// TIA Portal project "TESTV18" (V18) (continued)
REGION Network 8: HMI Command
   RUNG wire#powerrail
      Contact( "DB_AUX".HMI_Bit.HMIb5 )
      Coil( "DB_AUX".AXIS1.PLCToPCON.CTRL2.CTRL2_Sig_SON )
   END_RUNG
   RUNG wire#powerrail
      Contact( "DB_AUX".HMI_Bit.HMIb6 )
      Coil( "DB_AUX".AXIS1.PLCToPCON.CTRL2.CTRL2_Sig_DSTR )
   END_RUNG
   RUNG wire#powerrail
      Contact( "DB_AUX".HMI_Bit.HMIb7 )
      Coil( "DB_AUX".AXIS1.PLCToPCON.CTRL2.CTRL2_Sig_HOME )
   END_RUNG
   RUNG wire#powerrail
      Contact( "DB_AUX".HMI_Bit.HMIb8 )
      Coil( "DB_AUX".AXIS1.PLCToPCON.CTRL2."CTRL2_Sig_JOG+" )
   END_RUNG
   RUNG wire#powerrail
      Contact( "DB_AUX".HMI_Bit.HMIb9 )
      Coil( "DB_AUX".AXIS1.PLCToPCON.CTRL2."CTRL2_Sig_JOG-" )
   END_RUNG
   RUNG wire#powerrail
      Contact( "DB_AUX".HMI_Bit.HMIb10 )
      Coil( "DB_AUX".AXIS1.PLCToPCON.CTRL2.CTRL2_Sig_RES )
   END_RUNG
   // the same network as SCL:
   "DB_AUX".AXIS1.PLCToPCON.CTRL2.CTRL2_Sig_SON := "DB_AUX".HMI_Bit.HMIb5;
   "DB_AUX".AXIS1.PLCToPCON.CTRL2.CTRL2_Sig_DSTR := "DB_AUX".HMI_Bit.HMIb6;
   "DB_AUX".AXIS1.PLCToPCON.CTRL2.CTRL2_Sig_HOME := "DB_AUX".HMI_Bit.HMIb7;
   "DB_AUX".AXIS1.PLCToPCON.CTRL2."CTRL2_Sig_JOG+" := "DB_AUX".HMI_Bit.HMIb8;
   "DB_AUX".AXIS1.PLCToPCON.CTRL2."CTRL2_Sig_JOG-" := "DB_AUX".HMI_Bit.HMIb9;
   "DB_AUX".AXIS1.PLCToPCON.CTRL2.CTRL2_Sig_RES := "DB_AUX".HMI_Bit.HMIb10;
END_REGION
END_ORGANIZATION_BLOCK

// folder: LIBRERIE OPEN/0 Bit logic operations

FUNCTION "LGF_BitToggle" : DWord   // FC10033, SCL
TITLE = LGF_BitToggle
{ S7_Optimized_Access := 'TRUE' }
AUTHOR : Siemens_SIMATIC_Systems_Support
FAMILY : LGF
NAME : LGF_BitToggle
// Dieser Baustein toggelt (von TRUE nach FALSE und umgekehrt) ein Bit an vorgegebener Stelle in einer Variablen vom Datentyp DWORD.    
// Anstelle von DWord kann auch Word und Byte verwendet werden, indem der übergebene Parameter mit z. B. BYTE_TO_DWORD und das Ergebnis mit DWORD_TO_BYTE konvertiert wird.
// This block toggles (from TRUE to FALSE and vice versa) a bit at a predefined position in a variable of the data type DWORD.  
// Alternatively, Word and Byte can be used instead of DWord by converting the passed parameter with, for example, BYTE_TO_DWORD and the result with DWORD_TO_BYTE
   VAR_INPUT
      value : DWord;   // Tag where the bit has to be toggled / Variable, an der das Bit getoggelt wird.
      bitNo : USInt;   // Bit number to be toggled in the “value” parameter. / Bitnummer, die im Parameter "value" getoggelt werden soll.
   END_VAR
   // Ret_Val : Tag with toggled bit / Variable mit getoggeltem Bit.
   VAR CONSTANT
      TRUE_BOOL_BIT : DWord := 16#0001;   // Just one bit which is true, to shift in Dword for masking / Ein einzelnes Bit mit Wert := TRUE zum schieben im Dword und zur Maskierung
      MAX_NO_OF_BITS : USInt := 32;   // Maximum bits in a DWord = 32 / Maximalanzahl an Bits in einem Dword = 32
   END_VAR
BEGIN
   REGION BLOCK INFO HEADER
     //===============================================================================
     // SIEMENS AG / (c)Copyright 2019
     //-------------------------------------------------------------------------------
     // Title:            LGF_BitToggle
     // Comment/Function: Toggle bit in elementary datatype - DWord
     //                   can be used for Word and Byte as well, by convert
     //                   the passed paramter and the result using for e.g. Dword_to_Byte
     // Library/Family:   LGF (Library General Functions)
     // Author:           Siemens Digital Industry
     // Tested with:      CPU1212C DC/DC/DC FW:V4.2
     // Engineering:      TIA Portal V15.1
     // Restrictions:     ENO not in use, set to true, no error handling
     // Requirements:     PLC (S7-1200 / S7-1500)
     //-------------------------------------------------------------------------------
     // Change log table:
     // Version  | Date       | Expert in charge         | Changes applied
     // 01.00.00 | 06.06.2015 | Siemens Industry Support | first release
     // 03.00.00 | 23.04.2020 | Siemens Industry Support | Set version to V3.0.0
     //                         harmonize the version of the whole library
     // 03.00.01 | 19.01.2021 | Simatic Systems Support
     //                         Insert documentation
     //===============================================================================
   END_REGION

   REGION Logic
     // toggle the bit in tag
     // shift one true bit into given position
     // concatenate value then with XOR resets the bit on the given position
     #LGF_BitToggle := #value XOR SHL(IN := #TRUE_BOOL_BIT, N := (#bitNo MOD #MAX_NO_OF_BITS));

     // no error handling needed
     ENO := TRUE;
   END_REGION
END_FUNCTION

FUNCTION "LGF_BitSet" : DWord   // FC10078, SCL
TITLE = LGF_BitSet
{ S7_Optimized_Access := 'TRUE' }
AUTHOR : Siemens_SIMATIC_Systems_Support
FAMILY : LGF
NAME : LGF_BitSet
// Dieser Baustein setzt ein Bit an vorgegebener Stelle in einer Variable vom Daten-typ DWORD.  
// Anstelle von DWord kann auch Word und Byte verwendet werden, indem der übergebene Parameter mit z. B. BYTE_TO_DWORD und das Ergebnis mit DWORD_TO_BYTE konvertiert wird.
// This block sets a bit at a given position in a variable of the data type DWORD.  
// Alternatively, Word and Byte can be used instead of DWord by converting the passed parameter with, for example, BYTE_TO_DWORD and the result with DWORD_TO_BYTE.
   VAR_INPUT
      value : DWord;   // Tag where the bit has to be set / Variable, an der das Bit gesetzt wird
      bitNo : USInt;   // Bit number to set in "value" parameter / Bitnummer, die im Parameter "value" gesetzt werden soll
   END_VAR
   // Ret_Val : Tag with the set bit / Variable mit gesetztem Bit
   VAR CONSTANT
      TRUE_BOOL_BIT : DWord := 16#0001;   // Just one bit which is true, to shift in Dword for masking / Ein einzelnes Bit mit Wert := TRUE zum schieben im Dword und zur Maskierung
      MAX_NO_OF_BITS : USInt := 32;   // Maximum bits in a DWord = 32 / Maximalanzahl an Bits in einem Dword = 32
   END_VAR
BEGIN
   REGION BLOCK INFO HEADER
     //===============================================================================
     // SIEMENS AG / (c)Copyright 2019
     //-------------------------------------------------------------------------------
     // Title:            LGF_BitSet
     // Comment/Function: Set bit in elementary datatype - DWord
     //                   cam be used for Word and Byte as well, by convert
     //                   the passed paramter and the result using for e.g. Dword_to_Byte
     // Library/Family:   LGF (Library General Functions)
     // Author:           Siemens Digital Industry
     // Tested with:      CPU1212C DC/DC/DC FW:V4.2
     // Engineering:      TIA Portal V15.1
     // Restrictions:     ENO not in use, set to true, no error handling
     // Requirements:     PLC (S7-1200 / S7-1500)
     //-------------------------------------------------------------------------------
     // Change log table:
     // Version  | Date       | Expert in charge         | Changes applied
     // 01.00.00 | 06.06.2015 | Siemens Industry Support | first release
     // 03.00.00 | 23.04.2020 | Siemens Industry Support | Set version to V3.0.0
     //                         harmonize the version of the whole library
     // 03.00.01 | 19.01.2021 | Simatic Systems Support
     //                         Insert documentation
     //===============================================================================
   END_REGION

   REGION Logic
     // set the bit in tag
     // shift one true bit into given position
     // concatenate value then with OR will result in the previous value and the set bit in position
     #LGF_BitSet := #value OR SHL(IN := #TRUE_BOOL_BIT, N := (#bitNo MOD #MAX_NO_OF_BITS));

     // no error handling needed
     ENO := TRUE;
   END_REGION
END_FUNCTION

// folder: LIBRERIE OPEN/6 Converter operations/Binary types - Split and Merge

FUNCTION "LGF_MergeBitsToDWord" : DWord   // FC10062, SCL
TITLE = LGF_MergeBitsToDWord
{ S7_Optimized_Access := 'TRUE' }
AUTHOR : Siemens_Digital_Industry
FAMILY : LGF
NAME : LGF_MergeBitsToDWord
// This function merge 32 Bits / 32 Boolean variables into one DWord variable. / Diese Funktion führt 32 Bit / 32 Boolsche Variablen in einer DWord Variable zusammen.
   VAR_INPUT
      bit31 : Bool;   // Input Bit 31 - MSB
      bit30 : Bool;   // Input Bit 30
      bit29 : Bool;   // Input Bit 29
      bit28 : Bool;   // Input Bit 28
      bit27 : Bool;   // Input Bit 27
      bit26 : Bool;   // Input Bit 26
      bit25 : Bool;   // Input Bit 25
      bit24 : Bool;   // Input Bit 24
      bit23 : Bool;   // Input Bit 23
      bit22 : Bool;   // Input Bit 22
      bit21 : Bool;   // Input Bit 21
      bit20 : Bool;   // Input Bit 20
      bit19 : Bool;   // Input Bit 19
      bit18 : Bool;   // Input Bit 18
      bit17 : Bool;   // Input Bit 17
      bit16 : Bool;   // Input Bit 16
      bit15 : Bool;   // Input Bit 15
      bit14 : Bool;   // Input Bit 14
      bit13 : Bool;   // Input Bit 13
      bit12 : Bool;   // Input Bit 12
      bit11 : Bool;   // Input Bit 11
      bit10 : Bool;   // Input Bit 10
      bit9 : Bool;   // Input Bit 9
      bit8 : Bool;   // Input Bit 8
      bit7 : Bool;   // Input Bit 7
      bit6 : Bool;   // Input Bit 6
      bit5 : Bool;   // Input Bit 5
      bit4 : Bool;   // Input Bit 4
      bit3 : Bool;   // Input Bit 3
      bit2 : Bool;   // Input Bit 2
      bit1 : Bool;   // Input Bit 1
      bit0 : Bool;   // Input Bit 0 - LSB
   END_VAR
   VAR_TEMP
      tempDWord : DWord;   // Temp memory to merge Bits into a DWord / Temp speicher zum zusammenführen der Bits zu einem DWord
   END_VAR
   // Ret_Val : Composite Bit sequence stored as DWord variable / Zusammengefügte Bitfolge, gespeichert in einer DWord Variable
BEGIN
   REGION BLOCK INFO HEADER
     //===============================================================================
     // SIEMENS AG / (c)Copyright 2018
     //-------------------------------------------------------------------------------
     // Title:            LGF_MergeBitsToDWord
     // Comment/Function: This function merge 32 Bits / 32 Boolean variables into one DWord variable.
     // Library/Family:   LGF (Library General Functions)
     // Author:           Siemens Digital Industry Support
     // Tested with:      S7-PLCSIM Advanced V2.0 SP1
     // Engineering:      TIA Portal V14 / V14SP1
     // Restrictions:     ENO disabled - no error handling, no failure possible.
     // Requirements:     PLC (S7-1200 / S7-1500)
     //-------------------------------------------------------------------------------
     // Change log table:
     // Version  | Date       | Expert in charge       | Changes applied
     //----------|------------|------------------------|------------------------------
     // 01.00.00 | 20.06.2019 | Simatic Systems Support
     //                         First release
     // 03.00.00 | 23.04.2020 | Simatic Systems Support | Set version to V3.0.0
     //                         harmonize the version of the whole library
     // 03.00.01 | 22.02.2021 | Simatic Systems Support
     //                         Insert documentation
     //=============================================================================
   END_REGION

   REGION MERGE
     // set the bits by slice access
     #tempDWord.%X31 := #bit31;
     #tempDWord.%X30 := #bit30;
     #tempDWord.%X29 := #bit29;
     #tempDWord.%X28 := #bit28;
     #tempDWord.%X27 := #bit27;
     #tempDWord.%X26 := #bit26;
     #tempDWord.%X25 := #bit25;
     #tempDWord.%X24 := #bit24;
     #tempDWord.%X23 := #bit23;
     #tempDWord.%X22 := #bit22;
     #tempDWord.%X21 := #bit21;
     #tempDWord.%X20 := #bit20;
     #tempDWord.%X19 := #bit19;
     #tempDWord.%X18 := #bit18;
     #tempDWord.%X17 := #bit17;
     #tempDWord.%X16 := #bit16;
     #tempDWord.%X15 := #bit15;
     #tempDWord.%X14 := #bit14;
     #tempDWord.%X13 := #bit13;
     #tempDWord.%X12 := #bit12;
     #tempDWord.%X11 := #bit11;
     #tempDWord.%X10 := #bit10;
     #tempDWord.%X9 := #bit9;
     #tempDWord.%X8 := #bit8;
     #tempDWord.%X7 := #bit7;
     #tempDWord.%X6 := #bit6;
     #tempDWord.%X5 := #bit5;
     #tempDWord.%X4 := #bit4;
     #tempDWord.%X3 := #bit3;
     #tempDWord.%X2 := #bit2;
     #tempDWord.%X1 := #bit1;
     #tempDWord.%X0 := #bit0;
   END_REGION

   REGION OUTPUT
     #LGF_MergeBitsToDWord := #tempDWord;
     // no error handling needed
     ENO := TRUE;
   END_REGION
END_FUNCTION

FUNCTION "LGF_SplitDWordToBits" : Void   // FC10065, SCL
TITLE = LGF_SplitDWordToBits
{ S7_Optimized_Access := 'TRUE' }
AUTHOR : Siemens_Digital_Industry
FAMILY : LGF
NAME : LGF_SplitDWordToBits
// This function splits a DWord variable into 32 Boolean / 32 Bit variables. / Diese Funktion zerlegt eine DWord Variable in 32 Bool / 32 Bit Variablen.
   VAR_INPUT
      doubleWord : DWord;   // Bit sequence to be split / Bitfolge die zerlegt wird
   END_VAR
   VAR_OUTPUT
      bit31 : Bool;   // Output Bit 31 - MSB
      bit30 : Bool;   // Output Bit 30
      bit29 : Bool;   // Output Bit 29
      bit28 : Bool;   // Output Bit 28
      bit27 : Bool;   // Output Bit 27
      bit26 : Bool;   // Output Bit 26
      bit25 : Bool;   // Output Bit 25
      bit24 : Bool;   // Output Bit 24
      bit23 : Bool;   // Output Bit 23
      bit22 : Bool;   // Output Bit 22
      bit21 : Bool;   // Output Bit 21
      bit20 : Bool;   // Output Bit 20
      bit19 : Bool;   // Output Bit 19
      bit18 : Bool;   // Output Bit 18
      bit17 : Bool;   // Output Bit 17
      bit16 : Bool;   // Output Bit 16
      bit15 : Bool;   // Output Bit 15
      bit14 : Bool;   // Output Bit 14
      bit13 : Bool;   // Output Bit 13
      bit12 : Bool;   // Output Bit 12
      bit11 : Bool;   // Output Bit 11
      bit10 : Bool;   // Output Bit 10
      bit9 : Bool;   // Output Bit 9
      bit8 : Bool;   // Output Bit 8
      bit7 : Bool;   // Output Bit 7
      bit6 : Bool;   // Output Bit 6
      bit5 : Bool;   // Output Bit 5
      bit4 : Bool;   // Output Bit 4
      bit3 : Bool;   // Output Bit 3
      bit2 : Bool;   // Output Bit 2
      bit1 : Bool;   // Output Bit 1
      bit0 : Bool;   // Output Bit 0 - LSB
   END_VAR
BEGIN
   REGION BLOCK INFO HEADER
     //===============================================================================
     // SIEMENS AG / (c)Copyright 2018
     //-------------------------------------------------------------------------------
     // Title:            LGF_SplitDWordToBits
     // Comment/Function: This function splits a DWord variable into 32 Boolean / 32 Bit variables
     // Library/Family:   LGF (Library General Functions)
     // Author:           Siemens Digital Industry Support
     // Tested with:      S7-PLCSIM Advanced V2.0 SP1
     // Engineering:      TIA Portal V14 / V14SP1
     // Restrictions:     ENO disabled - no error handling, no failure possible.
     // Requirements:     PLC (S7-1200 / S7-1500)
     //-------------------------------------------------------------------------------
     // Change log table:
     // Version  | Date       | Expert in charge       | Changes applied
     //----------|------------|------------------------|------------------------------
     // 01.00.00 | 20.06.2019 | Simatic Systems Support
     //                         First release
     // 03.00.00 | 23.04.2020 | Simatic Systems Support | Set version to V3.0.0
     //                         harmonize the version of the whole library
     // 03.00.01 | 22.02.2021 | Simatic Systems Support
     //                         Insert documentation
     //=============================================================================
   END_REGION

   REGION OUTPUT
     // get the bits by slice access
     #bit31 := #doubleWord.%X31;
     #bit30 := #doubleWord.%X30;
     #bit29 := #doubleWord.%X29;
     #bit28 := #doubleWord.%X28;
     #bit27 := #doubleWord.%X27;
     #bit26 := #doubleWord.%X26;
     #bit25 := #doubleWord.%X25;
     #bit24 := #doubleWord.%X24;
     #bit23 := #doubleWord.%X23;
     #bit22 := #doubleWord.%X22;
     #bit21 := #doubleWord.%X21;
     #bit20 := #doubleWord.%X20;
     #bit19 := #doubleWord.%X19;
     #bit18 := #doubleWord.%X18;
     #bit17 := #doubleWord.%X17;
     #bit16 := #doubleWord.%X16;
     #bit15 := #doubleWord.%X15;
     #bit14 := #doubleWord.%X14;
     #bit13 := #doubleWord.%X13;
     #bit12 := #doubleWord.%X12;
     #bit11 := #doubleWord.%X11;
     #bit10 := #doubleWord.%X10;
     #bit9 := #doubleWord.%X9;
     #bit8 := #doubleWord.%X8;
     #bit7 := #doubleWord.%X7;
     #bit6 := #doubleWord.%X6;
     #bit5 := #doubleWord.%X5;
     #bit4 := #doubleWord.%X4;
     #bit3 := #doubleWord.%X3;
     #bit2 := #doubleWord.%X2;
     #bit1 := #doubleWord.%X1;
     #bit0 := #doubleWord.%X0;
     // no error handling needed
     ENO := TRUE;
   END_REGION
END_FUNCTION

// ===== library types =====

TYPE "Cylinder_Diagnostic"
   STRUCT
      Lost_Backward : Bool := FALSE;   // FC negativo perso / Negative HR verloren / Finecorsa indietro perso inaspettatamente
      Not_Reached_Backward : Bool := FALSE;   // FC negativo non raggiunto / Negative HR nicht erreicht / Finecorsa indietro non raggiunto
      Lost_Forward : Bool := FALSE;   // FC positivo perso / Positive HR verloren / Finecorsa avanti perso inaspettatamente
      Not_Reached_Forward : Bool := FALSE;   // FC positivo non raggiunto / Positive HR nicht erreicht / Finecorsa avanti non raggiunto
      Switch_Contemp : Bool := FALSE;   // FC negativo e positivo contemporanei / Gleichzeitige negative und positive HR / Finecorsa contemporanei
      Commands_Anomaly : Bool := FALSE;   // Comandi contemporanei / Zeitgenössische Befehle / Comandi contemporanei
   END_STRUCT;
END_TYPE

TYPE "Machine_Status_Data"
   STRUCT
      Power_On : Bool;   // Emergenze ok
      Power_On_Delayed : Bool;   // Emergenze ok con ritardo
      Pneumatic_On_Gen_Dly : Bool;   // Pneumatica generale OK
      AUTO_MODE : Bool;   // Modalità automatico
      MANU_MODE : Bool;   // Modalità manuale
      SBS_MODE : Bool;   // Modalità step by step
      End_Cycle_Request : Bool;   // Richiesta fine ciclo
      Empy_Pallet_Request : Bool;   // Richiesta svuotamento isola
      Alarm_Reset : Bool;   // Reset allarmi
      BarrieraImpegnata : Bool;   // Barriera Impegnata
      Bimano_OK : Bool;   // Bimanuale premuto
      Gen_alarm_ON : Bool;   // Allarme generale presente
      Gen_warn_ON : Bool;   // Warning generale presente
   END_STRUCT;
END_TYPE

// folder: Sensore digitale

TYPE "SENSOR_DIG"
TITLE = Sensor_DIG
// UDT per i dati di sensori digitali
   STRUCT
      Sensor_OUT : "Sensor_Dig_Out";   // Parametri d'uscita del sensore
      Sensor_PAR : "Sensor_Dig_Par";   // Parametri d'impostazione del sensore
   END_STRUCT;
END_TYPE

TYPE "Sensor_Dig_Out"
   STRUCT
      NO_Out : Bool;   // Uscita contatto diretto normalmente aperto / Normal open contact
      NC_Out : Bool;   // Uscita contatto diretto normalmente chiuso / Normal closed contact
      PE_Out : Bool;   // Uscita Fronte di salita segnale / Rising edge signal
      NE_Out : Bool;   // Uscita Fronte di discesa segnale / Falling edge signal
      OnDly_Out : Bool;   // Uscita con attivazione ritardata / Output delayed
      OffDly_Out : Bool;   // Uscita con isattivazione ritardata
   END_STRUCT;
END_TYPE

TYPE "Sensor_Dig_Par"
   STRUCT
      DLY_OnTime_S : IEC_TIMER;   // Temporizzatore per filtro lettura ON sensore / Delay timer filter ON sensor (S)
      DLY_OffTime_S : IEC_TIMER;   // Temporizzatore per filtro lettura OFF sensore / Delay timer filter OFF sensor (S)
      ME_PEOut : Bool;   // Memoria per appoggio fronte di salita / Positive edge flag
      ME_NEOut : Bool;   // Memoria per appoggio fronte di discesa
      TI_DlyOn_ms : Time;   // Valore tempo ritardo accensione ms / Timeout delay on S
      TI_DlyOff_ms : Time;   // Valore tempo ritardo spegnimento ms / Timeout delay off ms
   END_STRUCT;
END_TYPE

// folder: (top level)

FUNCTION_BLOCK "FB_AUTO_MANU_MODE"   // FB2, LAD
TITLE = FB_AUTO_MANU_MODE
{ S7_Optimized_Access := 'TRUE' }
AUTHOR : C.M.
VERSION : 0.1
// FB per la gestione delle modalità AUTO-MANU
   VAR_INPUT
      IV_AutoEnable : Bool;   // Ingresso abilitazione
      IV_AUX_INS_REQ : Bool;   // ingresso richiesta ausiliari
      IV_AUX_INSERTED : Bool;   // Ingresso ausiliari inseriti
      IV_AUTO_MODE_SEL : Bool;   // Ingresso selettore modale
      IV_START_CYCLE_BTN : Bool;   // Ingresso conferma attivazione modalità
      IV_END_CYCLE_BTN : Bool;   // Ingresso richiesta fine ciclo
      IV_END_CYCLE : Bool;   // Ingresso fine ciclo raggiunto
      IV_LAMP_TEST : Bool;   // Ingresso per test lampade
      IV_CLK_1Hz : Bool;   // Ingresso clock 1Hz
      IV_CLK_2Hz : Bool;   // Ingresso clock 2Hz
      IV_INFO : Bool;   // Ingresso lampada INFO
      IV_WARN : Bool;   // Ingresso lampada WARNING
      IV_ERROR : Bool;   // Ingresso lampada errore
   END_VAR
   VAR_OUTPUT
      OV_AUTO_MODE : Bool;   // Uscita modalità AUTO ON
      OV_MANU_MODE : Bool;   // Uscita modalità MANU ON
      OV_END_CYCLE_REQ : Bool;   // Uscita richiesta fine ciclo attivata
      OV_AUX_LAMP : Bool;   // Uscita per lampada ausiliari
      OV_CYCLE_LAMP : Bool;   // Uscita per lampada in ciclo
      OV_INFO_LAMP : Bool;   // Uscita per lampada info
      OV_WARN_LAMP : Bool;   // Uscita per lampada warning
      OV_ERROR_LAMP : Bool;   // Uscita per lampada errore
   END_VAR
   VAR
      ME_Mem1 : Bool;   // Memoria di appoggio AUTO ON
      FP_START_CYC_BTN : Bool;   // Appoggio fronte di salita start ciclo AUTO ON
      FP_END_CYC_STATUS : Bool;   // Appoggio fronte di salita richiesta fine ciclo
      R_TRIG1 : R_TRIG;   // Blocco fronte di salita 1
   END_VAR
   VAR_TEMP
      ME_EndCycleStatus : Bool;   // Memoria appoggio richiesta fine ciclo
   END_VAR
   VAR_TEMP   // added for the SCL form of the ladder/FBD networks
      _w1 : Bool;
      _w2 : Bool;
   END_VAR
BEGIN

REGION Network 1: Trigger start ciclo
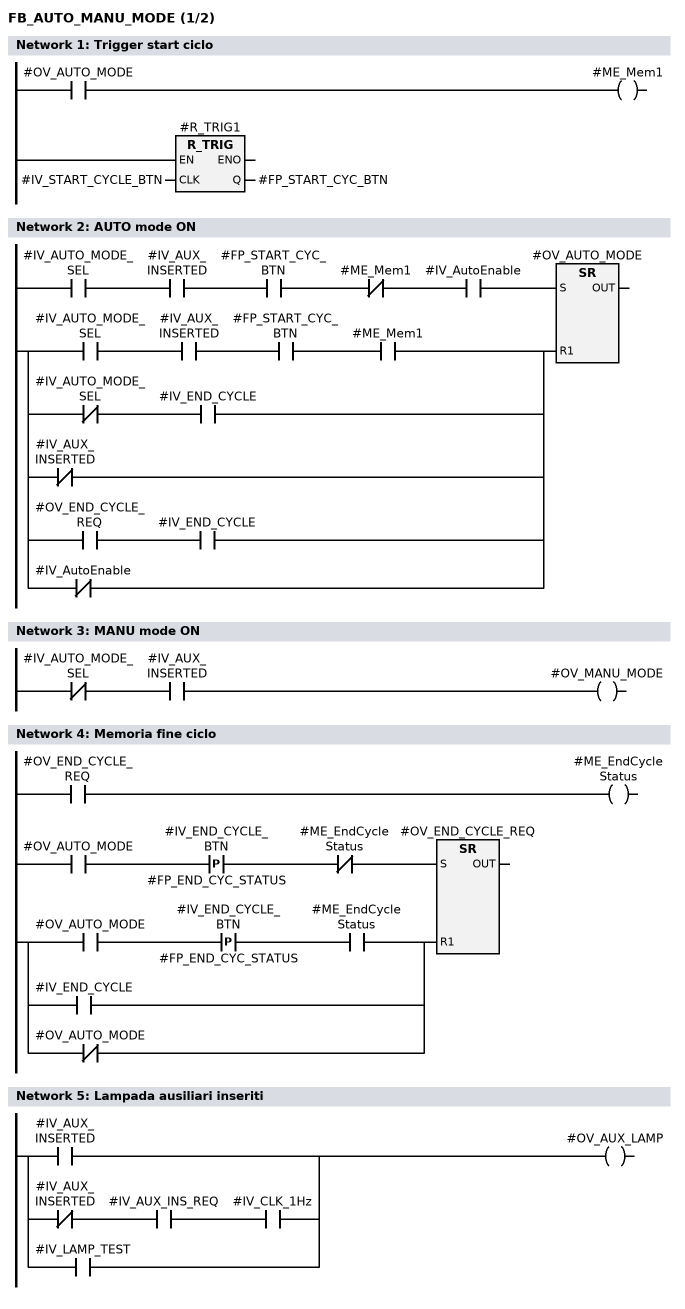
   #ME_Mem1 := #OV_AUTO_MODE;
   #R_TRIG1(CLK := #IV_START_CYCLE_BTN, Q => #FP_START_CYC_BTN);   // R_TRIG
END_REGION

REGION Network 2: AUTO mode ON
   RUNG wire#powerrail
      Contact( #IV_AUTO_MODE_SEL )
      Contact( #IV_AUX_INSERTED )
      Contact( #FP_START_CYC_BTN )
      I_Contact( #ME_Mem1 )
      Contact( #IV_AutoEnable )
      S_SR(operand := #OV_AUTO_MODE, r1 := wire#w1)
   END_RUNG
   RUNG wire#powerrail
      Contact( #IV_AUTO_MODE_SEL )
      Contact( #IV_AUX_INSERTED )
      Contact( #FP_START_CYC_BTN )
      Contact( #ME_Mem1 )
   END_RUNG wire#w1
   RUNG wire#powerrail
      I_Contact( #IV_AUTO_MODE_SEL )
      Contact( #IV_END_CYCLE )
   END_RUNG wire#w1
   RUNG wire#powerrail
      I_Contact( #IV_AUX_INSERTED )
   END_RUNG wire#w1
   RUNG wire#powerrail
      Contact( #OV_END_CYCLE_REQ )
      Contact( #IV_END_CYCLE )
   END_RUNG wire#w1
   RUNG wire#powerrail
      I_Contact( #IV_AutoEnable )
   END_RUNG wire#w1
   // the same network as SCL:
   IF #IV_AUTO_MODE_SEL AND #IV_AUX_INSERTED AND #FP_START_CYC_BTN AND NOT #ME_Mem1 AND #IV_AutoEnable THEN
       #OV_AUTO_MODE := TRUE;   // SR flip-flop
   END_IF;
   IF (#IV_AUTO_MODE_SEL AND #IV_AUX_INSERTED AND #FP_START_CYC_BTN AND #ME_Mem1) OR (NOT #IV_AUTO_MODE_SEL AND #IV_END_CYCLE) OR NOT #IV_AUX_INSERTED OR (#OV_END_CYCLE_REQ AND #IV_END_CYCLE) OR NOT #IV_AutoEnable THEN
       #OV_AUTO_MODE := FALSE;
   END_IF;
END_REGION

REGION Network 3: MANU mode ON
   RUNG wire#powerrail
      I_Contact( #IV_AUTO_MODE_SEL )
      Contact( #IV_AUX_INSERTED )
      Coil( #OV_MANU_MODE )
   END_RUNG
   // the same network as SCL:
   #OV_MANU_MODE := NOT #IV_AUTO_MODE_SEL AND #IV_AUX_INSERTED;
END_REGION

REGION Network 4: Memoria fine ciclo
   RUNG wire#powerrail
      Contact( #OV_END_CYCLE_REQ )
      Coil( #ME_EndCycleStatus )
   END_RUNG
   RUNG wire#powerrail
      Contact( #OV_AUTO_MODE )
      P_Contact(operand := #IV_END_CYCLE_BTN, bit := #FP_END_CYC_STATUS)
      I_Contact( #ME_EndCycleStatus )
      S_SR(operand := #OV_END_CYCLE_REQ, r1 := wire#w1)
   END_RUNG
   RUNG wire#powerrail
      Contact( #OV_AUTO_MODE )
      P_Contact(operand := #IV_END_CYCLE_BTN, bit := #FP_END_CYC_STATUS)
      Contact( #ME_EndCycleStatus )
   END_RUNG wire#w1
   RUNG wire#powerrail
      Contact( #IV_END_CYCLE )
   END_RUNG wire#w1
   RUNG wire#powerrail
      I_Contact( #OV_AUTO_MODE )
   END_RUNG wire#w1
   // the same network as SCL:
   #ME_EndCycleStatus := #OV_END_CYCLE_REQ;
   #_w1 := #OV_AUTO_MODE AND #IV_END_CYCLE_BTN AND NOT #FP_END_CYC_STATUS;   // rising edge of #IV_END_CYCLE_BTN
   #FP_END_CYC_STATUS := #IV_END_CYCLE_BTN;
   #_w2 := #OV_AUTO_MODE AND #IV_END_CYCLE_BTN AND NOT #FP_END_CYC_STATUS;   // rising edge of #IV_END_CYCLE_BTN
   #FP_END_CYC_STATUS := #IV_END_CYCLE_BTN;
   IF #_w1 AND NOT #ME_EndCycleStatus THEN
       #OV_END_CYCLE_REQ := TRUE;   // SR flip-flop
   END_IF;
   IF (#_w2 AND #ME_EndCycleStatus) OR #IV_END_CYCLE OR NOT #OV_AUTO_MODE THEN
       #OV_END_CYCLE_REQ := FALSE;
   END_IF;
END_REGION

REGION Network 5: Lampada ausiliari inseriti
   RUNG wire#powerrail
      Contact( #IV_AUX_INSERTED )
      wire#w1
      Coil( #OV_AUX_LAMP )
   END_RUNG
   RUNG wire#powerrail
      I_Contact( #IV_AUX_INSERTED )
      Contact( #IV_AUX_INS_REQ )
      Contact( #IV_CLK_1Hz )
   END_RUNG wire#w1
   RUNG wire#powerrail
      Contact( #IV_LAMP_TEST )
   END_RUNG wire#w1
   // the same network as SCL:
   #OV_AUX_LAMP := #IV_AUX_INSERTED OR (NOT #IV_AUX_INSERTED AND #IV_AUX_INS_REQ AND #IV_CLK_1Hz) OR #IV_LAMP_TEST;
END_REGION

REGION Network 6: Lampada in ciclo
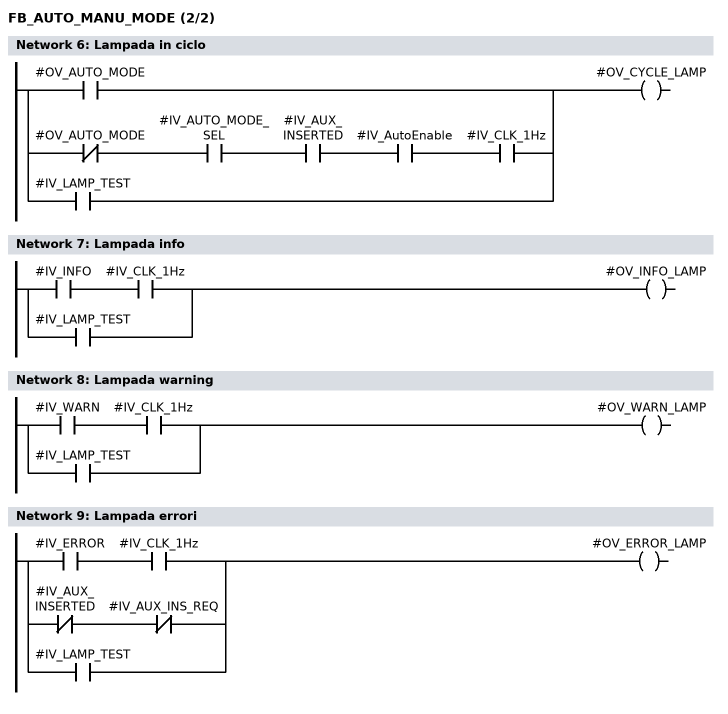
   RUNG wire#powerrail
      Contact( #OV_AUTO_MODE )
      wire#w1
      Coil( #OV_CYCLE_LAMP )
   END_RUNG
   RUNG wire#powerrail
      I_Contact( #OV_AUTO_MODE )
      Contact( #IV_AUTO_MODE_SEL )
      Contact( #IV_AUX_INSERTED )
      Contact( #IV_AutoEnable )
      Contact( #IV_CLK_1Hz )
   END_RUNG wire#w1
   RUNG wire#powerrail
      Contact( #IV_LAMP_TEST )
   END_RUNG wire#w1
   // the same network as SCL:
   #OV_CYCLE_LAMP := #OV_AUTO_MODE OR (NOT #OV_AUTO_MODE AND #IV_AUTO_MODE_SEL AND #IV_AUX_INSERTED AND #IV_AutoEnable AND #IV_CLK_1Hz) OR #IV_LAMP_TEST;
END_REGION

REGION Network 7: Lampada info
   RUNG wire#powerrail
      Contact( #IV_INFO )
      Contact( #IV_CLK_1Hz )
      wire#w1
      Coil( #OV_INFO_LAMP )
   END_RUNG
   RUNG wire#powerrail
      Contact( #IV_LAMP_TEST )
   END_RUNG wire#w1
   // the same network as SCL:
   #OV_INFO_LAMP := (#IV_INFO AND #IV_CLK_1Hz) OR #IV_LAMP_TEST;
END_REGION

REGION Network 8: Lampada warning
   RUNG wire#powerrail
      Contact( #IV_WARN )
      Contact( #IV_CLK_1Hz )
      wire#w1
      Coil( #OV_WARN_LAMP )
   END_RUNG
   RUNG wire#powerrail
      Contact( #IV_LAMP_TEST )
   END_RUNG wire#w1
   // the same network as SCL:
   #OV_WARN_LAMP := (#IV_WARN AND #IV_CLK_1Hz) OR #IV_LAMP_TEST;
END_REGION

REGION Network 9: Lampada errori
   RUNG wire#powerrail
      Contact( #IV_ERROR )
      Contact( #IV_CLK_1Hz )
      wire#w1
      Coil( #OV_ERROR_LAMP )
   END_RUNG
   RUNG wire#powerrail
      I_Contact( #IV_AUX_INSERTED )
      I_Contact( #IV_AUX_INS_REQ )
   END_RUNG wire#w1
   RUNG wire#powerrail
      Contact( #IV_LAMP_TEST )
   END_RUNG wire#w1
   // the same network as SCL:
   #OV_ERROR_LAMP := (#IV_ERROR AND #IV_CLK_1Hz) OR (NOT #IV_AUX_INSERTED AND NOT #IV_AUX_INS_REQ) OR #IV_LAMP_TEST;
END_REGION
END_FUNCTION_BLOCK

FUNCTION_BLOCK "FB_1WORD_GEN_ALLARMS"   // FB540, LAD
TITLE = FB_1W_GEN_ALLARMS
{ S7_Optimized_Access := 'TRUE' }
AUTHOR : C.M.
VERSION : 0.1
// FB per gestione di 1 word di allarmi
   VAR_INPUT
      IV_CND_ALLX0 : Bool;   // Ingresso per condizioni attivazione allarme X0
      IV_CND_ALLX1 : Bool;   // Ingresso per condizioni attivazione allarme X1
      IV_CND_ALLX2 : Bool;   // Ingresso per condizioni attivazione allarme X2
      IV_CND_ALLX3 : Bool;   // Ingresso per condizioni attivazione allarme X3
      IV_CND_ALLX4 : Bool;   // Ingresso per condizioni attivazione allarme X4
      IV_CND_ALLX5 : Bool;   // Ingresso per condizioni attivazione allarme X5
      IV_CND_ALLX6 : Bool;   // Ingresso per condizioni attivazione allarme X6
      IV_CND_ALLX7 : Bool;   // Ingresso per condizioni attivazione allarme X7
      IV_CND_ALLX8 : Bool;   // Ingresso per condizioni attivazione allarme X8
      IV_CND_ALLX9 : Bool;   // Ingresso per condizioni attivazione allarme X9
      IV_CND_ALLX10 : Bool;   // Ingresso per condizioni attivazione allarme X10
      IV_CND_ALLX11 : Bool;   // Ingresso per condizioni attivazione allarme X11
      IV_CND_ALLX12 : Bool;   // Ingresso per condizioni attivazione allarme X12
      IV_CND_ALLX13 : Bool;   // Ingresso per condizioni attivazione allarme X13
      IV_CND_ALLX14 : Bool;   // Ingresso per condizioni attivazione allarme X14
      IV_CND_ALLX15 : Bool;   // Ingresso per condizioni attivazione allarme X15
      IV_RST_ALL : Bool;   // Ingresso per RESET allarmi
   END_VAR
   VAR_OUTPUT
      VW_Allarms : Word;   // Variabile di uscita WORD per allarmi
   END_VAR
   VAR
      TI_T0 : IEC_TIMER;   // Timer attivazione allarme bit X0
      TI_T1 : IEC_TIMER;   // Timer attivazione allarme bit X1
      TI_T2 : IEC_TIMER;   // Timer attivazione allarme bit X2
      TI_T3 : IEC_TIMER;   // Timer attivazione allarme bit X3
      TI_T4 : IEC_TIMER;   // Timer attivazione allarme bit X4
      TI_T5 : IEC_TIMER;   // Timer attivazione allarme bit X5
      TI_T6 : IEC_TIMER;   // Timer attivazione allarme bit X6
      TI_T7 : IEC_TIMER;   // Timer attivazione allarme bit X7
      TI_T8 : IEC_TIMER;   // Timer attivazione allarme bit X8
      TI_T9 : IEC_TIMER;   // Timer attivazione allarme bit X9
      TI_T10 : IEC_TIMER;   // Timer attivazione allarme bit X10
      TI_T11 : IEC_TIMER;   // Timer attivazione allarme bit X11
      TI_T12 : IEC_TIMER;   // Timer attivazione allarme bit X12
      TI_T13 : IEC_TIMER;   // Timer attivazione allarme bit X13
      TI_T14 : IEC_TIMER;   // Timer attivazione allarme bit X14
      TI_T15 : IEC_TIMER;   // Timer attivazione allarme bit X15
   END_VAR
   VAR_TEMP   // added for the SCL form of the ladder/FBD networks
      _w1 : Bool;
   END_VAR
   // TI_T0.PT := T#5s;
   // TI_T1.PT := T#5s;
   // TI_T2.PT := T#5s;
   // TI_T3.PT := T#5s;
   // TI_T4.PT := T#5s;
   // TI_T5.PT := T#5s;
   // TI_T6.PT := T#5s;
   // TI_T7.PT := T#5s;
   // TI_T8.PT := T#5s;
   // TI_T9.PT := T#5s;
   // TI_T10.PT := T#5s;
   // TI_T11.PT := T#5s;
   // TI_T12.PT := T#5s;
   // TI_T13.PT := T#5s;
   // TI_T14.PT := T#5s;
   // TI_T15.PT := T#5s;
BEGIN

REGION Network 1: Bit X0 = Allarme 1
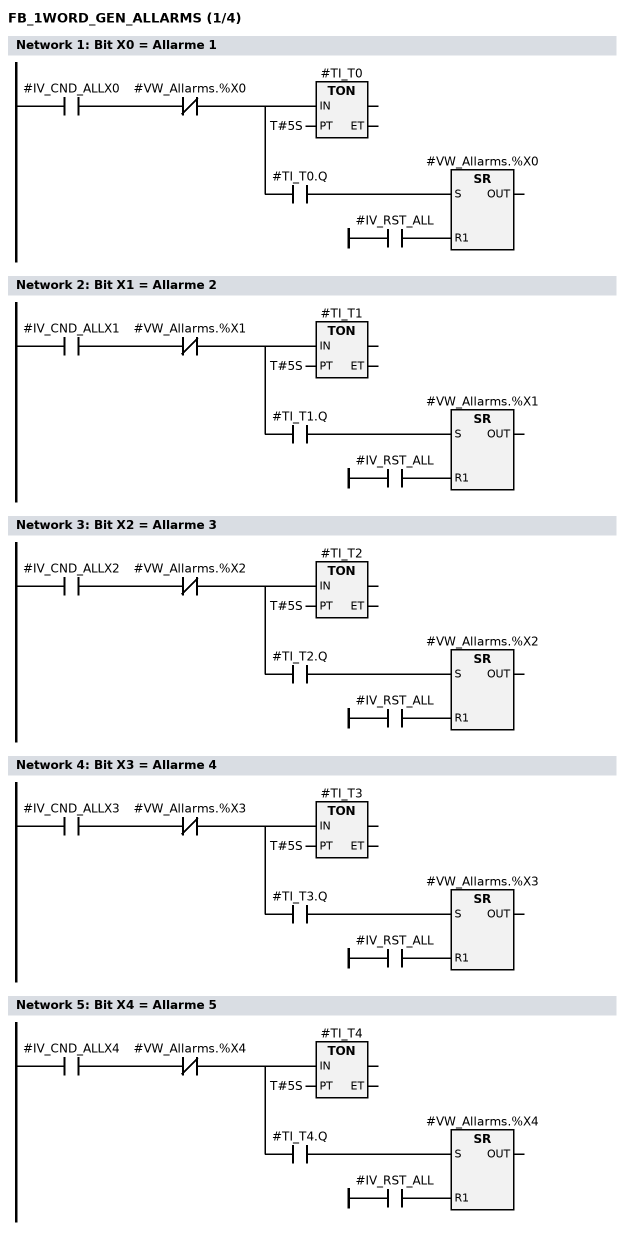
   #_w1 := #IV_CND_ALLX0 AND NOT #VW_Allarms.%X0;
   #TI_T0.TON(IN := #_w1, PT := T#5S);
   IF #_w1 AND #TI_T0.Q THEN
       #VW_Allarms.%X0 := TRUE;   // SR flip-flop
   END_IF;
   IF #IV_RST_ALL THEN #VW_Allarms.%X0 := FALSE; END_IF;
END_REGION

REGION Network 2: Bit X1 = Allarme 2
   #_w1 := #IV_CND_ALLX1 AND NOT #VW_Allarms.%X1;
   #TI_T1.TON(IN := #_w1, PT := T#5S);
   IF #_w1 AND #TI_T1.Q THEN
       #VW_Allarms.%X1 := TRUE;   // SR flip-flop
   END_IF;
   IF #IV_RST_ALL THEN #VW_Allarms.%X1 := FALSE; END_IF;
END_REGION

REGION Network 3: Bit X2 = Allarme 3
   #_w1 := #IV_CND_ALLX2 AND NOT #VW_Allarms.%X2;
   #TI_T2.TON(IN := #_w1, PT := T#5S);
   IF #_w1 AND #TI_T2.Q THEN
       #VW_Allarms.%X2 := TRUE;   // SR flip-flop
   END_IF;
   IF #IV_RST_ALL THEN #VW_Allarms.%X2 := FALSE; END_IF;
END_REGION

REGION Network 4: Bit X3 = Allarme 4
   #_w1 := #IV_CND_ALLX3 AND NOT #VW_Allarms.%X3;
   #TI_T3.TON(IN := #_w1, PT := T#5S);
   IF #_w1 AND #TI_T3.Q THEN
       #VW_Allarms.%X3 := TRUE;   // SR flip-flop
   END_IF;
   IF #IV_RST_ALL THEN #VW_Allarms.%X3 := FALSE; END_IF;
END_REGION

REGION Network 5: Bit X4 = Allarme 5
   #_w1 := #IV_CND_ALLX4 AND NOT #VW_Allarms.%X4;
   #TI_T4.TON(IN := #_w1, PT := T#5S);
   IF #_w1 AND #TI_T4.Q THEN
       #VW_Allarms.%X4 := TRUE;   // SR flip-flop
   END_IF;
   IF #IV_RST_ALL THEN #VW_Allarms.%X4 := FALSE; END_IF;
END_REGION

REGION Network 6: Bit X5 = Allarme 6
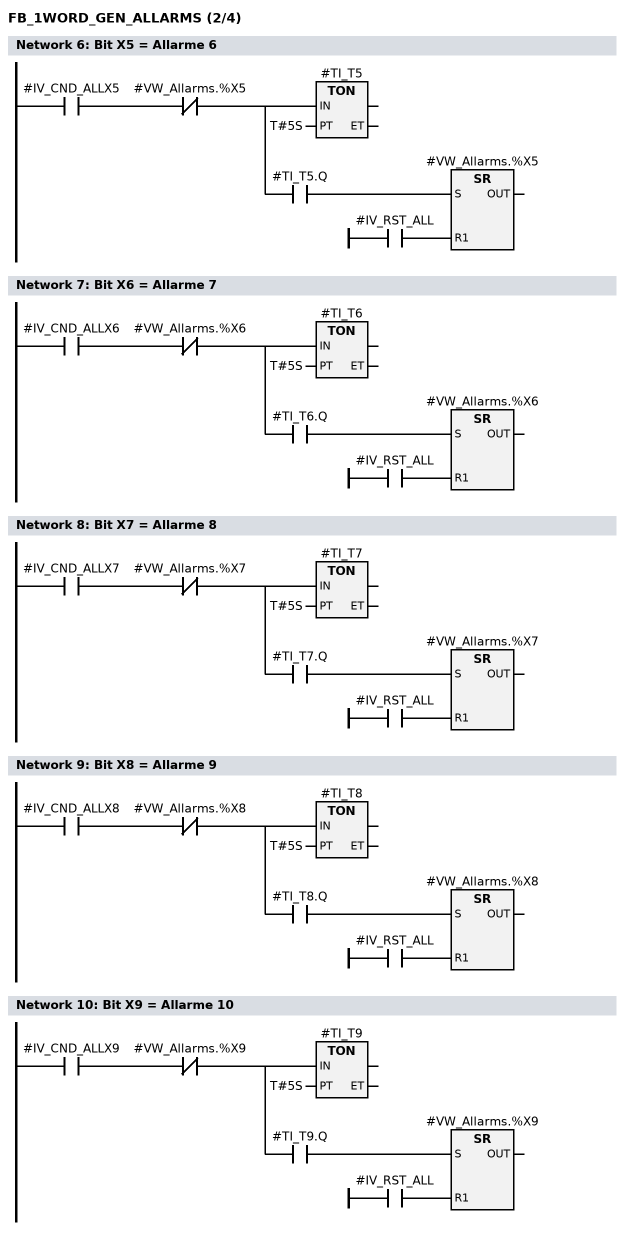
   #_w1 := #IV_CND_ALLX5 AND NOT #VW_Allarms.%X5;
   #TI_T5.TON(IN := #_w1, PT := T#5S);
   IF #_w1 AND #TI_T5.Q THEN
       #VW_Allarms.%X5 := TRUE;   // SR flip-flop
   END_IF;
   IF #IV_RST_ALL THEN #VW_Allarms.%X5 := FALSE; END_IF;
END_REGION

REGION Network 7: Bit X6 = Allarme 7
   #_w1 := #IV_CND_ALLX6 AND NOT #VW_Allarms.%X6;
   #TI_T6.TON(IN := #_w1, PT := T#5S);
   IF #_w1 AND #TI_T6.Q THEN
       #VW_Allarms.%X6 := TRUE;   // SR flip-flop
   END_IF;
   IF #IV_RST_ALL THEN #VW_Allarms.%X6 := FALSE; END_IF;
END_REGION

REGION Network 8: Bit X7 = Allarme 8
   #_w1 := #IV_CND_ALLX7 AND NOT #VW_Allarms.%X7;
   #TI_T7.TON(IN := #_w1, PT := T#5S);
   IF #_w1 AND #TI_T7.Q THEN
       #VW_Allarms.%X7 := TRUE;   // SR flip-flop
   END_IF;
   IF #IV_RST_ALL THEN #VW_Allarms.%X7 := FALSE; END_IF;
END_REGION

REGION Network 9: Bit X8 = Allarme 9
   #_w1 := #IV_CND_ALLX8 AND NOT #VW_Allarms.%X8;
   #TI_T8.TON(IN := #_w1, PT := T#5S);
   IF #_w1 AND #TI_T8.Q THEN
       #VW_Allarms.%X8 := TRUE;   // SR flip-flop
   END_IF;
   IF #IV_RST_ALL THEN #VW_Allarms.%X8 := FALSE; END_IF;
END_REGION

REGION Network 10: Bit X9 = Allarme 10
   #_w1 := #IV_CND_ALLX9 AND NOT #VW_Allarms.%X9;
   #TI_T9.TON(IN := #_w1, PT := T#5S);
   IF #_w1 AND #TI_T9.Q THEN
       #VW_Allarms.%X9 := TRUE;   // SR flip-flop
   END_IF;
   IF #IV_RST_ALL THEN #VW_Allarms.%X9 := FALSE; END_IF;
END_REGION

REGION Network 11: Bit X10 = Allarme 11
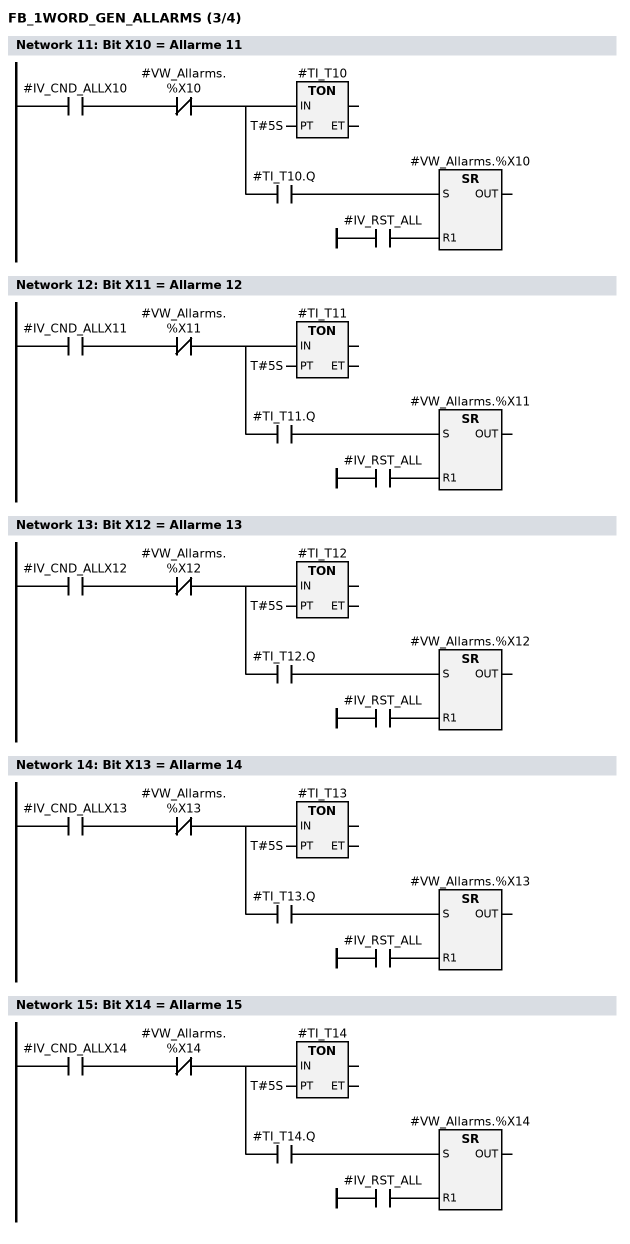
   #_w1 := #IV_CND_ALLX10 AND NOT #VW_Allarms.%X10;
   #TI_T10.TON(IN := #_w1, PT := T#5S);
   IF #_w1 AND #TI_T10.Q THEN
       #VW_Allarms.%X10 := TRUE;   // SR flip-flop
   END_IF;
   IF #IV_RST_ALL THEN #VW_Allarms.%X10 := FALSE; END_IF;
END_REGION

REGION Network 12: Bit X11 = Allarme 12
   #_w1 := #IV_CND_ALLX11 AND NOT #VW_Allarms.%X11;
   #TI_T11.TON(IN := #_w1, PT := T#5S);
   IF #_w1 AND #TI_T11.Q THEN
       #VW_Allarms.%X11 := TRUE;   // SR flip-flop
   END_IF;
   IF #IV_RST_ALL THEN #VW_Allarms.%X11 := FALSE; END_IF;
END_REGION
